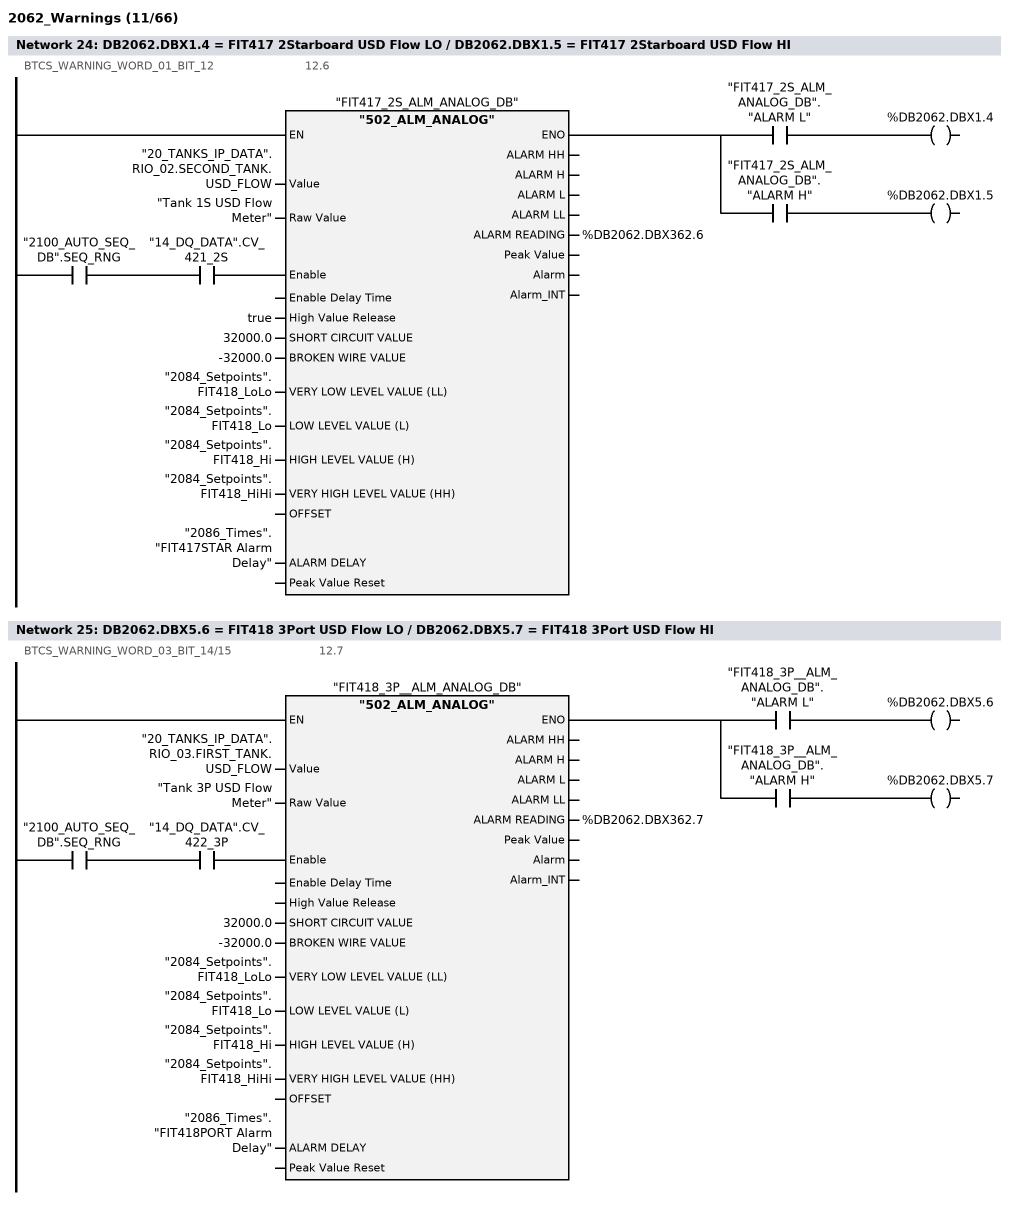
   RUNG wire#powerrail
      "FIT417_2S_ALM_ANALOG_DB"(Enable := wire#w1, Value := "20_TANKS_IP_DATA".RIO_02.SECOND_TANK.USD_FLOW, "Raw Value" := "Tank 1S USD Flow Meter", "Enable Delay Time" :=, "High Value Release" := true, "SHORT CIRCUIT VALUE" := 32000.0, "BROKEN WIRE VALUE" := -32000.0, "VERY LOW LEVEL VALUE (LL)" := "2084_Setpoints".FIT418_LoLo, "LOW LEVEL VALUE (L)" := "2084_Setpoints".FIT418_Lo, "HIGH LEVEL VALUE (H)" := "2084_Setpoints".FIT418_Hi, "VERY HIGH LEVEL VALUE (HH)" := "2084_Setpoints".FIT418_HiHi, OFFSET :=, "ALARM DELAY" := "2086_Times"."FIT417STAR Alarm Delay", "Peak Value Reset" :=, "ALARM HH" =>, "ALARM H" =>, "ALARM L" =>, "ALARM LL" =>, "ALARM READING" => %DB2062.DBX362.6, "Peak Value" =>, Alarm =>, Alarm_INT =>)
      wire#w2
      Contact( "FIT417_2S_ALM_ANALOG_DB"."ALARM L" )
      Coil( %DB2062.DBX1.4 )
   END_RUNG
   RUNG wire#powerrail
      Contact( "2100_AUTO_SEQ_DB".SEQ_RNG )
      Contact( "14_DQ_DATA".CV_421_2S )
   END_RUNG wire#w1
   RUNG wire#w2
      Contact( "FIT417_2S_ALM_ANALOG_DB"."ALARM H" )
      Coil( %DB2062.DBX1.5 )
   END_RUNG
   // the same network as SCL:
   "FIT417_2S_ALM_ANALOG_DB"(Value := "20_TANKS_IP_DATA".RIO_02.SECOND_TANK.USD_FLOW,   // "502_ALM_ANALOG"
                           "Raw Value" := "Tank 1S USD Flow Meter",
                           Enable := "2100_AUTO_SEQ_DB".SEQ_RNG AND "14_DQ_DATA".CV_421_2S,
                           "High Value Release" := true,
                           "SHORT CIRCUIT VALUE" := 32000.0,
                           "BROKEN WIRE VALUE" := -32000.0,
                           "VERY LOW LEVEL VALUE (LL)" := "2084_Setpoints".FIT418_LoLo,
                           "LOW LEVEL VALUE (L)" := "2084_Setpoints".FIT418_Lo,
                           "HIGH LEVEL VALUE (H)" := "2084_Setpoints".FIT418_Hi,
                           "VERY HIGH LEVEL VALUE (HH)" := "2084_Setpoints".FIT418_HiHi,
                           "ALARM DELAY" := "2086_Times"."FIT417STAR Alarm Delay",
                           "ALARM READING" => %DB2062.DBX362.6,
                           ENO => #_w1);
   %DB2062.DBX1.4 := #_w1 AND "FIT417_2S_ALM_ANALOG_DB"."ALARM L";
   %DB2062.DBX1.5 := #_w1 AND "FIT417_2S_ALM_ANALOG_DB"."ALARM H";
END_REGION

REGION Network 25: DB2062.DBX5.6 = FIT418 3Port USD Flow LO / DB2062.DBX5.7 = FIT418 3Port USD Flow HI
   // BTCS_WARNING_WORD_03_BIT_14/15                         12.7
   RUNG wire#powerrail
      "FIT418_3P__ALM_ANALOG_DB"(Enable := wire#w1, Value := "20_TANKS_IP_DATA".RIO_03.FIRST_TANK.USD_FLOW, "Raw Value" := "Tank 3P USD Flow Meter", "Enable Delay Time" :=, "High Value Release" :=, "SHORT CIRCUIT VALUE" := 32000.0, "BROKEN WIRE VALUE" := -32000.0, "VERY LOW LEVEL VALUE (LL)" := "2084_Setpoints".FIT418_LoLo, "LOW LEVEL VALUE (L)" := "2084_Setpoints".FIT418_Lo, "HIGH LEVEL VALUE (H)" := "2084_Setpoints".FIT418_Hi, "VERY HIGH LEVEL VALUE (HH)" := "2084_Setpoints".FIT418_HiHi, OFFSET :=, "ALARM DELAY" := "2086_Times"."FIT418PORT Alarm Delay", "Peak Value Reset" :=, "ALARM HH" =>, "ALARM H" =>, "ALARM L" =>, "ALARM LL" =>, "ALARM READING" => %DB2062.DBX362.7, "Peak Value" =>, Alarm =>, Alarm_INT =>)
      wire#w2
      Contact( "FIT418_3P__ALM_ANALOG_DB"."ALARM L" )
      Coil( %DB2062.DBX5.6 )
   END_RUNG
   RUNG wire#powerrail
      Contact( "2100_AUTO_SEQ_DB".SEQ_RNG )
      Contact( "14_DQ_DATA".CV_422_3P )
   END_RUNG wire#w1
   RUNG wire#w2
      Contact( "FIT418_3P__ALM_ANALOG_DB"."ALARM H" )
      Coil( %DB2062.DBX5.7 )
   END_RUNG
   // the same network as SCL:
   "FIT418_3P__ALM_ANALOG_DB"(Value := "20_TANKS_IP_DATA".RIO_03.FIRST_TANK.USD_FLOW,   // "502_ALM_ANALOG"
                           "Raw Value" := "Tank 3P USD Flow Meter",
                           Enable := "2100_AUTO_SEQ_DB".SEQ_RNG AND "14_DQ_DATA".CV_422_3P,
                           "SHORT CIRCUIT VALUE" := 32000.0,
                           "BROKEN WIRE VALUE" := -32000.0,
                           "VERY LOW LEVEL VALUE (LL)" := "2084_Setpoints".FIT418_LoLo,
                           "LOW LEVEL VALUE (L)" := "2084_Setpoints".FIT418_Lo,
                           "HIGH LEVEL VALUE (H)" := "2084_Setpoints".FIT418_Hi,
                           "VERY HIGH LEVEL VALUE (HH)" := "2084_Setpoints".FIT418_HiHi,
                           "ALARM DELAY" := "2086_Times"."FIT418PORT Alarm Delay",
                           "ALARM READING" => %DB2062.DBX362.7,
                           ENO => #_w1);
   %DB2062.DBX5.6 := #_w1 AND "FIT418_3P__ALM_ANALOG_DB"."ALARM L";
   %DB2062.DBX5.7 := #_w1 AND "FIT418_3P__ALM_ANALOG_DB"."ALARM H";
END_REGION

REGION Network 26: DB2062.DBX6.0 = FIT417 3Starboard USD Flow LO / DB2062.DBX6.1 = FIT417 3Starboard USD Flow HI
   // BTCS_WARNING_WORD_04_BIT_0/1                              12.8
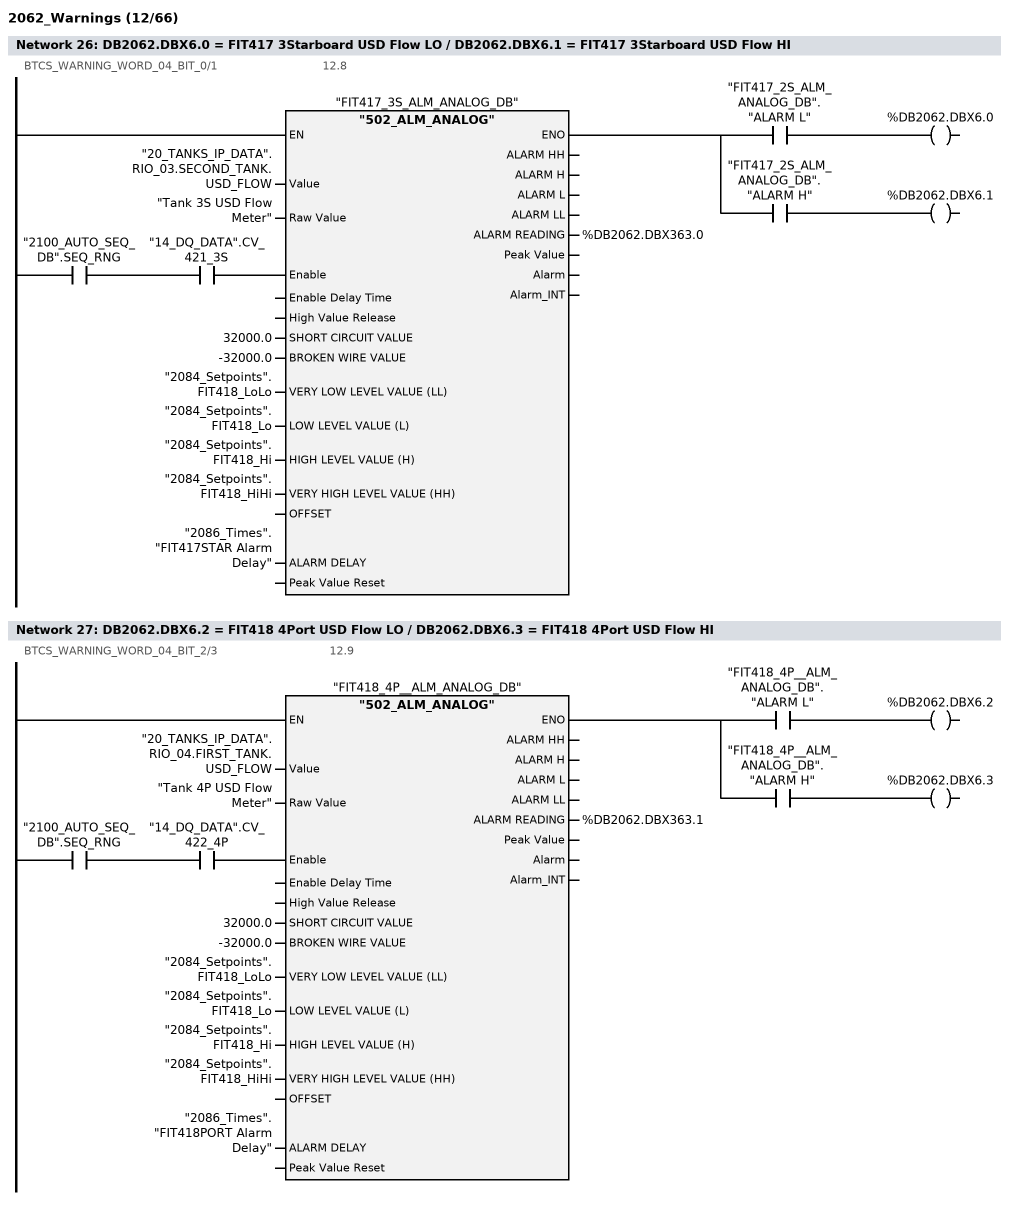
   RUNG wire#powerrail
      "FIT417_3S_ALM_ANALOG_DB"(Enable := wire#w1, Value := "20_TANKS_IP_DATA".RIO_03.SECOND_TANK.USD_FLOW, "Raw Value" := "Tank 3S USD Flow Meter", "Enable Delay Time" :=, "High Value Release" :=, "SHORT CIRCUIT VALUE" := 32000.0, "BROKEN WIRE VALUE" := -32000.0, "VERY LOW LEVEL VALUE (LL)" := "2084_Setpoints".FIT418_LoLo, "LOW LEVEL VALUE (L)" := "2084_Setpoints".FIT418_Lo, "HIGH LEVEL VALUE (H)" := "2084_Setpoints".FIT418_Hi, "VERY HIGH LEVEL VALUE (HH)" := "2084_Setpoints".FIT418_HiHi, OFFSET :=, "ALARM DELAY" := "2086_Times"."FIT417STAR Alarm Delay", "Peak Value Reset" :=, "ALARM HH" =>, "ALARM H" =>, "ALARM L" =>, "ALARM LL" =>, "ALARM READING" => %DB2062.DBX363.0, "Peak Value" =>, Alarm =>, Alarm_INT =>)
      wire#w2
      Contact( "FIT417_2S_ALM_ANALOG_DB"."ALARM L" )
      Coil( %DB2062.DBX6.0 )
   END_RUNG
   RUNG wire#powerrail
      Contact( "2100_AUTO_SEQ_DB".SEQ_RNG )
      Contact( "14_DQ_DATA".CV_421_3S )
   END_RUNG wire#w1
   RUNG wire#w2
      Contact( "FIT417_2S_ALM_ANALOG_DB"."ALARM H" )
      Coil( %DB2062.DBX6.1 )
   END_RUNG
   // the same network as SCL:
   "FIT417_3S_ALM_ANALOG_DB"(Value := "20_TANKS_IP_DATA".RIO_03.SECOND_TANK.USD_FLOW,   // "502_ALM_ANALOG"
                           "Raw Value" := "Tank 3S USD Flow Meter",
                           Enable := "2100_AUTO_SEQ_DB".SEQ_RNG AND "14_DQ_DATA".CV_421_3S,
                           "SHORT CIRCUIT VALUE" := 32000.0,
                           "BROKEN WIRE VALUE" := -32000.0,
                           "VERY LOW LEVEL VALUE (LL)" := "2084_Setpoints".FIT418_LoLo,
                           "LOW LEVEL VALUE (L)" := "2084_Setpoints".FIT418_Lo,
                           "HIGH LEVEL VALUE (H)" := "2084_Setpoints".FIT418_Hi,
                           "VERY HIGH LEVEL VALUE (HH)" := "2084_Setpoints".FIT418_HiHi,
                           "ALARM DELAY" := "2086_Times"."FIT417STAR Alarm Delay",
                           "ALARM READING" => %DB2062.DBX363.0,
                           ENO => #_w1);
   %DB2062.DBX6.0 := #_w1 AND "FIT417_2S_ALM_ANALOG_DB"."ALARM L";
   %DB2062.DBX6.1 := #_w1 AND "FIT417_2S_ALM_ANALOG_DB"."ALARM H";
END_REGION

REGION Network 27: DB2062.DBX6.2 = FIT418 4Port USD Flow LO / DB2062.DBX6.3 = FIT418 4Port USD Flow HI
   // BTCS_WARNING_WORD_04_BIT_2/3                                12.9
   RUNG wire#powerrail
      "FIT418_4P__ALM_ANALOG_DB"(Enable := wire#w1, Value := "20_TANKS_IP_DATA".RIO_04.FIRST_TANK.USD_FLOW, "Raw Value" := "Tank 4P USD Flow Meter", "Enable Delay Time" :=, "High Value Release" :=, "SHORT CIRCUIT VALUE" := 32000.0, "BROKEN WIRE VALUE" := -32000.0, "VERY LOW LEVEL VALUE (LL)" := "2084_Setpoints".FIT418_LoLo, "LOW LEVEL VALUE (L)" := "2084_Setpoints".FIT418_Lo, "HIGH LEVEL VALUE (H)" := "2084_Setpoints".FIT418_Hi, "VERY HIGH LEVEL VALUE (HH)" := "2084_Setpoints".FIT418_HiHi, OFFSET :=, "ALARM DELAY" := "2086_Times"."FIT418PORT Alarm Delay", "Peak Value Reset" :=, "ALARM HH" =>, "ALARM H" =>, "ALARM L" =>, "ALARM LL" =>, "ALARM READING" => %DB2062.DBX363.1, "Peak Value" =>, Alarm =>, Alarm_INT =>)
      wire#w2
      Contact( "FIT418_4P__ALM_ANALOG_DB"."ALARM L" )
      Coil( %DB2062.DBX6.2 )
   END_RUNG
   RUNG wire#powerrail
      Contact( "2100_AUTO_SEQ_DB".SEQ_RNG )
      Contact( "14_DQ_DATA".CV_422_4P )
   END_RUNG wire#w1
   RUNG wire#w2
      Contact( "FIT418_4P__ALM_ANALOG_DB"."ALARM H" )
      Coil( %DB2062.DBX6.3 )
   END_RUNG
   // the same network as SCL:
   "FIT418_4P__ALM_ANALOG_DB"(Value := "20_TANKS_IP_DATA".RIO_04.FIRST_TANK.USD_FLOW,   // "502_ALM_ANALOG"
                           "Raw Value" := "Tank 4P USD Flow Meter",
                           Enable := "2100_AUTO_SEQ_DB".SEQ_RNG AND "14_DQ_DATA".CV_422_4P,
                           "SHORT CIRCUIT VALUE" := 32000.0,
                           "BROKEN WIRE VALUE" := -32000.0,
                           "VERY LOW LEVEL VALUE (LL)" := "2084_Setpoints".FIT418_LoLo,
                           "LOW LEVEL VALUE (L)" := "2084_Setpoints".FIT418_Lo,
                           "HIGH LEVEL VALUE (H)" := "2084_Setpoints".FIT418_Hi,
                           "VERY HIGH LEVEL VALUE (HH)" := "2084_Setpoints".FIT418_HiHi,
                           "ALARM DELAY" := "2086_Times"."FIT418PORT Alarm Delay",
                           "ALARM READING" => %DB2062.DBX363.1,
                           ENO => #_w1);
   %DB2062.DBX6.2 := #_w1 AND "FIT418_4P__ALM_ANALOG_DB"."ALARM L";
   %DB2062.DBX6.3 := #_w1 AND "FIT418_4P__ALM_ANALOG_DB"."ALARM H";
END_REGION

REGION Network 28: DB2062.DBX6.4 = FIT417 4Starboard USD Flow LO / DB2062.DBX6.5 = FIT417 4Starboard USD Flow HI
   // BTCS_WARNING_WORD_04_BIT_4/5                        12.10
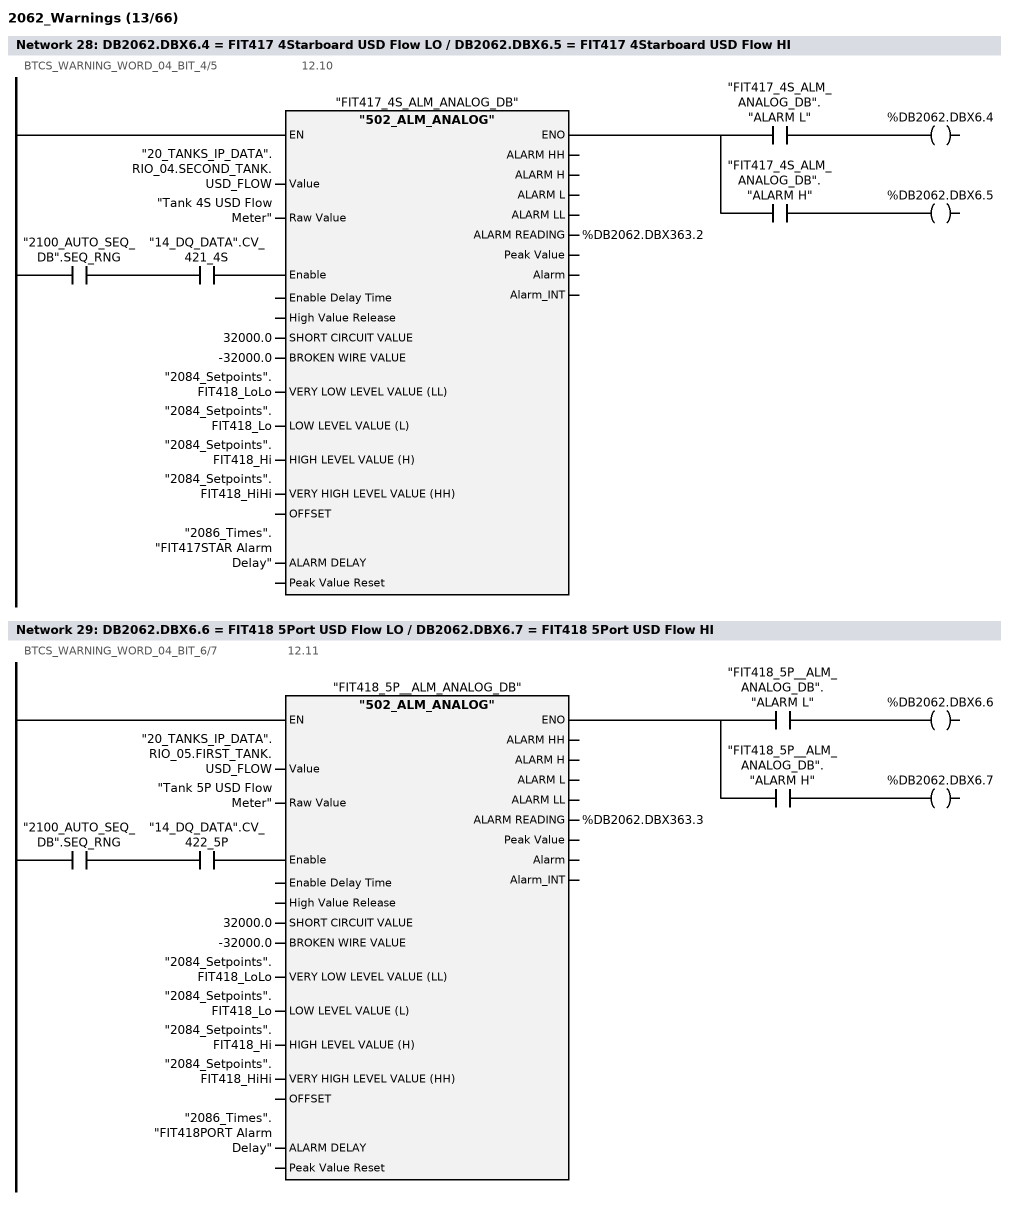
   RUNG wire#powerrail
      "FIT417_4S_ALM_ANALOG_DB"(Enable := wire#w1, Value := "20_TANKS_IP_DATA".RIO_04.SECOND_TANK.USD_FLOW, "Raw Value" := "Tank 4S USD Flow Meter", "Enable Delay Time" :=, "High Value Release" :=, "SHORT CIRCUIT VALUE" := 32000.0, "BROKEN WIRE VALUE" := -32000.0, "VERY LOW LEVEL VALUE (LL)" := "2084_Setpoints".FIT418_LoLo, "LOW LEVEL VALUE (L)" := "2084_Setpoints".FIT418_Lo, "HIGH LEVEL VALUE (H)" := "2084_Setpoints".FIT418_Hi, "VERY HIGH LEVEL VALUE (HH)" := "2084_Setpoints".FIT418_HiHi, OFFSET :=, "ALARM DELAY" := "2086_Times"."FIT417STAR Alarm Delay", "Peak Value Reset" :=, "ALARM HH" =>, "ALARM H" =>, "ALARM L" =>, "ALARM LL" =>, "ALARM READING" => %DB2062.DBX363.2, "Peak Value" =>, Alarm =>, Alarm_INT =>)
      wire#w2
      Contact( "FIT417_4S_ALM_ANALOG_DB"."ALARM L" )
      Coil( %DB2062.DBX6.4 )
   END_RUNG
   RUNG wire#powerrail
      Contact( "2100_AUTO_SEQ_DB".SEQ_RNG )
      Contact( "14_DQ_DATA".CV_421_4S )
   END_RUNG wire#w1
   RUNG wire#w2
      Contact( "FIT417_4S_ALM_ANALOG_DB"."ALARM H" )
      Coil( %DB2062.DBX6.5 )
   END_RUNG
   // the same network as SCL:
   "FIT417_4S_ALM_ANALOG_DB"(Value := "20_TANKS_IP_DATA".RIO_04.SECOND_TANK.USD_FLOW,   // "502_ALM_ANALOG"
                           "Raw Value" := "Tank 4S USD Flow Meter",
                           Enable := "2100_AUTO_SEQ_DB".SEQ_RNG AND "14_DQ_DATA".CV_421_4S,
                           "SHORT CIRCUIT VALUE" := 32000.0,
                           "BROKEN WIRE VALUE" := -32000.0,
                           "VERY LOW LEVEL VALUE (LL)" := "2084_Setpoints".FIT418_LoLo,
                           "LOW LEVEL VALUE (L)" := "2084_Setpoints".FIT418_Lo,
                           "HIGH LEVEL VALUE (H)" := "2084_Setpoints".FIT418_Hi,
                           "VERY HIGH LEVEL VALUE (HH)" := "2084_Setpoints".FIT418_HiHi,
                           "ALARM DELAY" := "2086_Times"."FIT417STAR Alarm Delay",
                           "ALARM READING" => %DB2062.DBX363.2,
                           ENO => #_w1);
   %DB2062.DBX6.4 := #_w1 AND "FIT417_4S_ALM_ANALOG_DB"."ALARM L";
   %DB2062.DBX6.5 := #_w1 AND "FIT417_4S_ALM_ANALOG_DB"."ALARM H";
END_REGION

REGION Network 29: DB2062.DBX6.6 = FIT418 5Port USD Flow LO / DB2062.DBX6.7 = FIT418 5Port USD Flow HI
   // BTCS_WARNING_WORD_04_BIT_6/7                    12.11
   RUNG wire#powerrail
      "FIT418_5P__ALM_ANALOG_DB"(Enable := wire#w1, Value := "20_TANKS_IP_DATA".RIO_05.FIRST_TANK.USD_FLOW, "Raw Value" := "Tank 5P USD Flow Meter", "Enable Delay Time" :=, "High Value Release" :=, "SHORT CIRCUIT VALUE" := 32000.0, "BROKEN WIRE VALUE" := -32000.0, "VERY LOW LEVEL VALUE (LL)" := "2084_Setpoints".FIT418_LoLo, "LOW LEVEL VALUE (L)" := "2084_Setpoints".FIT418_Lo, "HIGH LEVEL VALUE (H)" := "2084_Setpoints".FIT418_Hi, "VERY HIGH LEVEL VALUE (HH)" := "2084_Setpoints".FIT418_HiHi, OFFSET :=, "ALARM DELAY" := "2086_Times"."FIT418PORT Alarm Delay", "Peak Value Reset" :=, "ALARM HH" =>, "ALARM H" =>, "ALARM L" =>, "ALARM LL" =>, "ALARM READING" => %DB2062.DBX363.3, "Peak Value" =>, Alarm =>, Alarm_INT =>)
      wire#w2
      Contact( "FIT418_5P__ALM_ANALOG_DB"."ALARM L" )
      Coil( %DB2062.DBX6.6 )
   END_RUNG
   RUNG wire#powerrail
      Contact( "2100_AUTO_SEQ_DB".SEQ_RNG )
      Contact( "14_DQ_DATA".CV_422_5P )
   END_RUNG wire#w1
   RUNG wire#w2
      Contact( "FIT418_5P__ALM_ANALOG_DB"."ALARM H" )
      Coil( %DB2062.DBX6.7 )
   END_RUNG
   // the same network as SCL:
   "FIT418_5P__ALM_ANALOG_DB"(Value := "20_TANKS_IP_DATA".RIO_05.FIRST_TANK.USD_FLOW,   // "502_ALM_ANALOG"
                           "Raw Value" := "Tank 5P USD Flow Meter",
                           Enable := "2100_AUTO_SEQ_DB".SEQ_RNG AND "14_DQ_DATA".CV_422_5P,
                           "SHORT CIRCUIT VALUE" := 32000.0,
                           "BROKEN WIRE VALUE" := -32000.0,
                           "VERY LOW LEVEL VALUE (LL)" := "2084_Setpoints".FIT418_LoLo,
                           "LOW LEVEL VALUE (L)" := "2084_Setpoints".FIT418_Lo,
                           "HIGH LEVEL VALUE (H)" := "2084_Setpoints".FIT418_Hi,
                           "VERY HIGH LEVEL VALUE (HH)" := "2084_Setpoints".FIT418_HiHi,
                           "ALARM DELAY" := "2086_Times"."FIT418PORT Alarm Delay",
                           "ALARM READING" => %DB2062.DBX363.3,
                           ENO => #_w1);
   %DB2062.DBX6.6 := #_w1 AND "FIT418_5P__ALM_ANALOG_DB"."ALARM L";
   %DB2062.DBX6.7 := #_w1 AND "FIT418_5P__ALM_ANALOG_DB"."ALARM H";
END_REGION

REGION Network 30: DB2062.DBX7.0 = FIT417 5Starboard USD Flow LO / DB2062.DBX7.1 = FIT417 5Starboard USD Flow HI
   // BTCS_WARNING_WORD_04_BIT_8/9                         12.12
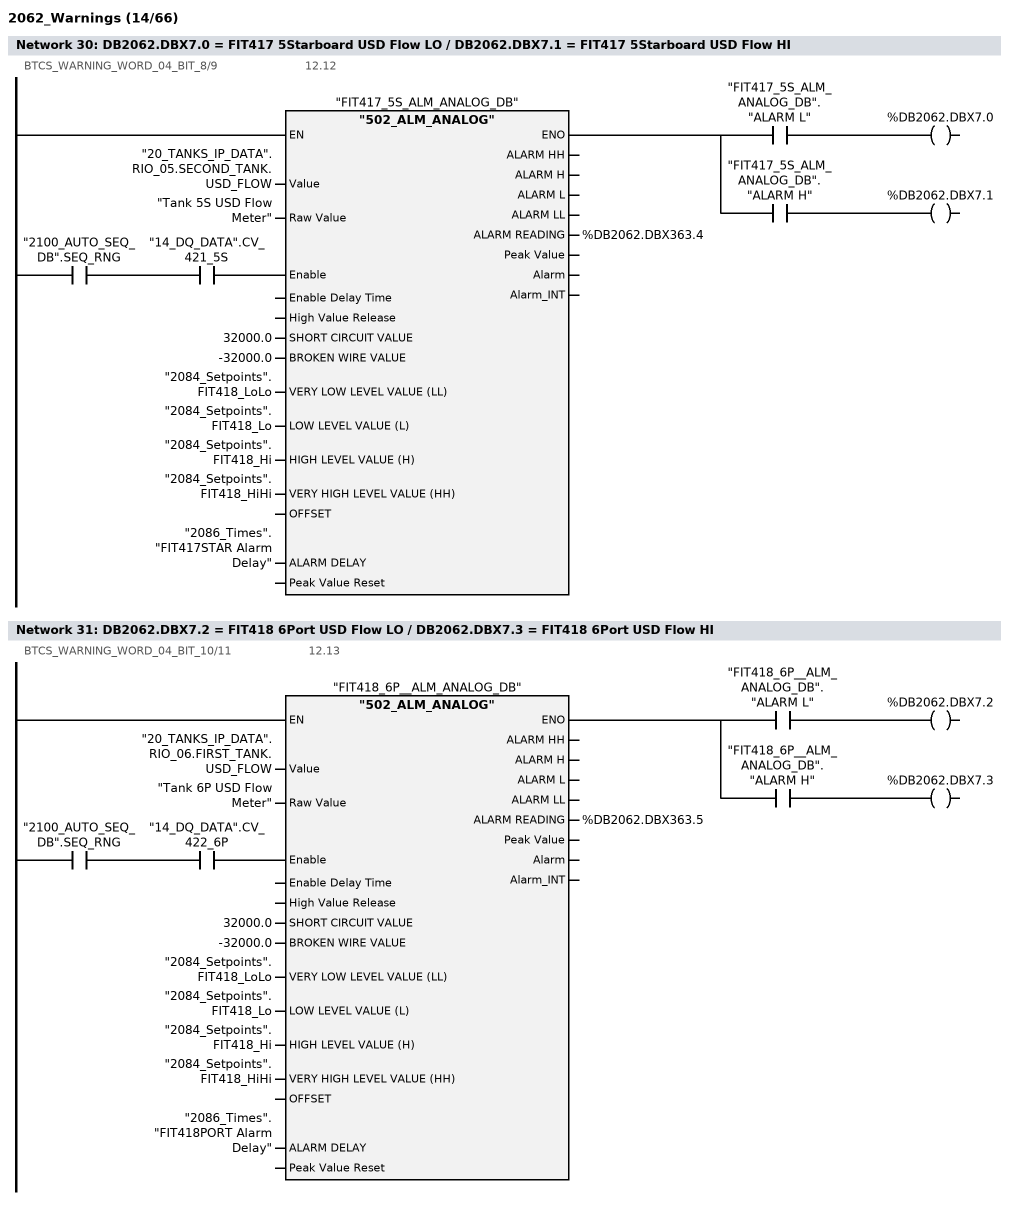
   RUNG wire#powerrail
      "FIT417_5S_ALM_ANALOG_DB"(Enable := wire#w1, Value := "20_TANKS_IP_DATA".RIO_05.SECOND_TANK.USD_FLOW, "Raw Value" := "Tank 5S USD Flow Meter", "Enable Delay Time" :=, "High Value Release" :=, "SHORT CIRCUIT VALUE" := 32000.0, "BROKEN WIRE VALUE" := -32000.0, "VERY LOW LEVEL VALUE (LL)" := "2084_Setpoints".FIT418_LoLo, "LOW LEVEL VALUE (L)" := "2084_Setpoints".FIT418_Lo, "HIGH LEVEL VALUE (H)" := "2084_Setpoints".FIT418_Hi, "VERY HIGH LEVEL VALUE (HH)" := "2084_Setpoints".FIT418_HiHi, OFFSET :=, "ALARM DELAY" := "2086_Times"."FIT417STAR Alarm Delay", "Peak Value Reset" :=, "ALARM HH" =>, "ALARM H" =>, "ALARM L" =>, "ALARM LL" =>, "ALARM READING" => %DB2062.DBX363.4, "Peak Value" =>, Alarm =>, Alarm_INT =>)
      wire#w2
      Contact( "FIT417_5S_ALM_ANALOG_DB"."ALARM L" )
      Coil( %DB2062.DBX7.0 )
   END_RUNG
   RUNG wire#powerrail
      Contact( "2100_AUTO_SEQ_DB".SEQ_RNG )